   12662: 'Pump6: Pressure recording: warning, value undershot', class Pump Warning Alarm, trigger "Pump6_Pressure_Record_DBW_142" bit 10
   12663: 'Pump6: Pressure recording: fault, value exceeded', class Pump Error Alarm, trigger "Pump6_Pressure_Record_DBW_142" bit 11
   12664: 'Pump6: Pressure recording: fault, value undershot', class Pump Error Alarm, trigger "Pump6_Pressure_Record_DBW_142" bit 12
   12665: 'Pump6: Temp. recording HP heat exch.: measured value outside measuring range', class Pump Warning Alarm, trigger "Pump6_Heatexchanger_DBW_220" bit 8
   12666: 'Pump6: Temp. recording HP heat exch.: warning, value exceeded', class Pump Warning Alarm, trigger "Pump6_Heatexchanger_DBW_220" bit 9
   12667: 'Pump6: Temp. recording HP heat exch.: warning, value undershot', class Pump Warning Alarm, trigger "Pump6_Heatexchanger_DBW_220" bit 10
   12668: 'Pump6: Temp. recording HP heat exch.: fault, value exceeded', class Pump Error Alarm, trigger "Pump6_Heatexchanger_DBW_220" bit 11
   12669: 'Pump6: Temp. recording HP heat exch.: fault, value undershot', class Pump Error Alarm, trigger "Pump6_Heatexchanger_DBW_220" bit 12
   10101: 'Mixinghead hydraulic: Motor protection switch has tripped', class Mixing Hydraulic Errors, trigger "Mixinghead_Hydraulic_DBW2" bit 8
   10102: 'Mixinghead hydraulic: Min. fill level hydraulic oil undershot', class Mixing Hydraulic Errors, trigger "Mixinghead_Hydraulic_DBW2" bit 9
   10103: 'Mixinghead hydraulic: Warning max. temperature exceeded', class Mixing Hydraulic Warning, trigger "Mixinghead_Hydraulic_DBW2" bit 10
   10104: 'Mixinghead hydraulic: HP filter contaminated', class Mixing Hydraulic Warning, trigger "Mixinghead_Hydraulic_DBW2" bit 11
   10105: 'Mixinghead hydraulic: Activation max. temperature exceeded', class Mixing Hydraulic Errors, trigger "Mixinghead_Hydraulic_DBW2" bit 12
   10106: 'Mixinghead hydraulic: Return filter contaminated', class Mixing Hydraulic Warning, trigger "Mixinghead_Hydraulic_DBW2" bit 13
   10107: 'Mixinghead hydraulic: Cable break at pressure switch', class Mixing Hydraulic Errors, trigger "Mixinghead_Hydraulic_DBW2" bit 14
   10108: 'Mixinghead hydraulic: Max. pressure not reached', class Mixing Hydraulic Errors, trigger "Mixinghead_Hydraulic_DBW2" bit 15
   10109: 'Mixinghead hydraulic: Moog filter contaminated', class Mixing Hydraulic Warning, trigger "Mixinghead_Hydraulic_DBW2" bit 0
   10110: 'Mixinghead hydraulic: Min. fill level filter pump', class Mixing Hydraulic Warning, trigger "Mixinghead_Hydraulic_DBW2" bit 1
   10111: 'Mixinghead hydraulic: Motor protecting switch of filter pump tripped', class Mixing Hydraulic Errors, trigger "Mixinghead_Hydraulic_DBW2" bit 2
   10112: 'Mixinghead hydraulic: Max. fill level filter pump', class Mixing Hydraulic Errors, trigger "Mixinghead_Hydraulic_DBW2" bit 3
   10113: 'Mixinghead hydraulic: Filter bypass fault', class Mixing Hydraulic Warning, trigger "Mixinghead_Hydraulic_DBW2" bit 4
   10114: 'Mixinghead hydraulic:', class Mixing Hydraulic Warning, trigger "Mixinghead_Hydraulic_DBW2" bit 5
   10115: 'Mixinghead hydraulic:', class Mixing Hydraulic Errors, trigger "Mixinghead_Hydraulic_DBW2" bit 6
   10116: 'Mixinghead hydraulic:', class Mixing Hydraulic Errors, trigger "Mixinghead_Hydraulic_DBW2" bit 7
   15001: 'Mixinghead 01: Mixinghead does not open', class Mixing Head Errors, trigger "Mixinghead_MHControl1_DBW_2" bit 8
   15002: 'Mixinghead 01: Mixinghead does not close', class Mixing Head Errors, trigger "Mixinghead_MHControl1_DBW_2" bit 9
   15003: 'Mixinghead 01: Entry cancelled', class Mixing Head Warning, trigger "Mixinghead_MHControl1_DBW_2" bit 10
   15004: 'Mixinghead 01: Mixinghead open without activation', class Mixing Head Errors, trigger "Mixinghead_MHControl1_DBW_2" bit 11
   15005: 'Mixinghead 01: Mixinghead close during entry', class Mixing Head Warning, trigger "Mixinghead_MHControl1_DBW_2" bit 12
   15006: 'Mixinghead 01: Warning, shot time too short', class Mixing Head Warning, trigger "Mixinghead_MHControl1_DBW_2" bit 13
   15007: 'Mixinghead 01: Warning , shot time too long', class Mixing Head Warning, trigger "Mixinghead_MHControl1_DBW_2" bit 14
   15008: 'Mixinghead 01: Fault, shot time too short', class Mixing Head Warning, trigger "Mixinghead_MHControl1_DBW_2" bit 15
   15009: 'Mixinghead 01: Mixinghead collides when opening or closing', class Mixing Head Warning, trigger "Mixinghead_MHControl1_DBW_2" bit 0
   15010: 'Mixinghead 01: Runtime monitoring when locking mixing head', class Mixing Head Warning, trigger "Mixinghead_MHControl1_DBW_2" bit 1
   15011: 'Mixinghead 01: Runtime monitoring when unlocking mixing head', class Mixing Head Warning, trigger "Mixinghead_MHControl1_DBW_2" bit 2
   15012: 'Mixinghead 01:', class Mixing Head Warning, trigger "Mixinghead_MHControl1_DBW_2" bit 3
   15013: 'Mixinghead 01: Min. Pressure for the cleaning air', class Mixing Head Warning, trigger "Mixinghead_MHControl1_DBW_2" bit 4
   15014: 'Mixinghead 01: Max. Pressure for the cleaning air', class Mixing Head Warning, trigger "Mixinghead_MHControl1_DBW_2" bit 5
   15015: 'Mixinghead 01:', class Mixing Head Warning, trigger "Mixinghead_MHControl1_DBW_2" bit 6
   15016: 'Mixinghead 01: Component required in entry is not enabled at this mixing head', class Mixing Head Errors, trigger "Mixinghead_MHControl1_DBW_2" bit 7
   15017: 'Mixinghead 01: Cleaning piston: Moving out too slow', class Mixing Head Errors, trigger "Mixinghead_Cpiston1_DBW_34" bit 8
   15018: 'Mixinghead 01: Cleaning piston: Moving in too slow', class Mixing Head Errors, trigger "Mixinghead_Cpiston1_DBW_34" bit 9
   15019: 'Mixinghead 01: Cleaning piston: Proximity switch defect', class Mixinghead Error Archive Foaming, trigger "Mixinghead_Cpiston1_DBW_34" bit 10
   15020: 'Mixinghead 01: Cleaning piston: Leaves its home position in entry', class Mixing Head Errors, trigger "Mixinghead_Cpiston1_DBW_34" bit 11
   15021: 'Mixinghead 01: Cleaning piston: Not defined', class Mixing Head Warning, trigger "Mixinghead_Cpiston1_DBW_34" bit 12
   15022: 'Mixinghead 01: Cleaning piston:', class Mixing Head Warning, trigger "Mixinghead_Cpiston1_DBW_34" bit 13
   15023: 'Mixinghead 01: Cleaning piston:', class Mixing Head Warning, trigger "Mixinghead_Cpiston1_DBW_34" bit 14
   15024: 'Mixinghead 01: Cleaning piston:', class Mixing Head Warning, trigger "Mixinghead_Cpiston1_DBW_34" bit 15
   15025: 'Mixinghead 01: Cleaning piston: Controller at upper limit', class Mixing Head Warning, trigger "Mixinghead_Cpiston1_DBW_34" bit 0
   15026: 'Mixinghead 01: Cleaning piston: Controller at lower limit', class Mixing Head Warning, trigger "Mixinghead_Cpiston1_DBW_34" bit 1
   15027: 'Mixinghead 01: Cleaning piston:', class Mixing Head Warning, trigger "Mixinghead_Cpiston1_DBW_34" bit 2
   15028: 'Mixinghead 01: Cleaning piston: Front position not reached', class Mixing Head Warning, trigger "Mixinghead_Cpiston1_DBW_34" bit 3
   15029: 'Mixinghead 01: Cleaning piston: Rear position not reached', class Mixing Head Warning, trigger "Mixinghead_Cpiston1_DBW_34" bit 4
   15030: 'Mixinghead 01: Cleaning piston: Home position not reached', class Mixing Head Warning, trigger "Mixinghead_Cpiston1_DBW_34" bit 5
   15031: 'Mixinghead 01: Cleaning piston:', class Mixing Head Warning, trigger "Mixinghead_Cpiston1_DBW_34" bit 6
   15032: 'Mixinghead 01: Cleaning piston:', class Mixing Head Warning, trigger "Mixinghead_Cpiston1_DBW_34" bit 7
   15040: 'Mixinghead 01: Connection 01: Temperature recording: Measuring value outside measuring range', class Mixinghead Warn Archv Foam, trigger "Mixinghead_Temperature_MH1_Con1_DBW70" bit 8
   15041: 'Mixinghead 01: Connection 01: Temperature recording: Warning, value exceeded', class Mixing Head Warning, trigger "Mixinghead_Temperature_MH1_Con1_DBW70" bit 9
   15042: 'Mixinghead 01: Connection 01: Temperature recording: Warning, value undershot', class Mixing Head Warning, trigger "Mixinghead_Temperature_MH1_Con1_DBW70" bit 10
   15043: 'Mixinghead 01: Connection 01: Temperature recording: Fault, value exceeded', class Mixing Head Errors, trigger "Mixinghead_Temperature_MH1_Con1_DBW70" bit 11
   15044: 'Mixinghead 01: Connection 01: Temperature recording: Fault, value undershot', class Mixing Head Errors, trigger "Mixinghead_Temperature_MH1_Con1_DBW70" bit 12
   15045: 'Mixinghead 01: Connection 02: Temperature recording: Measuring value outside measuring range', class Mixinghead Warn Archv Foam, trigger "Mixinghead_Temperature_MH1_Con2_DBW104" bit 8
   15046: 'Mixinghead 01: Connection 02: Temperature recording: Warning, value exceeded', class Mixing Head Warning, trigger "Mixinghead_Temperature_MH1_Con2_DBW104" bit 9
   15047: 'Mixinghead 01: Connection 02: Temperature recording: Warning, value undershot', class Mixing Head Warning, trigger "Mixinghead_Temperature_MH1_Con2_DBW104" bit 10
   15048: 'Mixinghead 01: Connection 02: Temperature recording: Fault, value exceeded', class Mixing Head Errors, trigger "Mixinghead_Temperature_MH1_Con2_DBW104" bit 11
   15049: 'Mixinghead 01: Connection 02: Temperature recording: Fault, value undershot', class Mixing Head Errors, trigger "Mixinghead_Temperature_MH1_Con2_DBW104" bit 12
   15050: 'Mixinghead 01: Connection 03: Temperature recording: Measuring value outside measuring range', class Mixing Head Warning, trigger "Mixinghead_Temperature_MH1_Con3_DBW138" bit 8
   15051: 'Mixinghead 01: Connection 03: Temperature recording: Warning, value exceeded', class Mixing Head Warning, trigger "Mixinghead_Temperature_MH1_Con3_DBW138" bit 9
   15052: 'Mixinghead 01: Connection 03: Temperature recording: Warning, value undershot', class Mixing Head Warning, trigger "Mixinghead_Temperature_MH1_Con3_DBW138" bit 10
   15053: 'Mixinghead 01: Connection 03: Temperature recording: Fault, value exceeded', class Mixing Head Errors, trigger "Mixinghead_Temperature_MH1_Con3_DBW138" bit 11
   15054: 'Mixinghead 01: Connection 03: Temperature recording: Fault, value undershot', class Mixing Head Errors, trigger "Mixinghead_Temperature_MH1_Con3_DBW138" bit 12
   15055: 'Mixinghead 01: Connection 04: Temperature recording: Measuring value outside measuring range', class Mixing Head Warning, trigger "Mixinghead_Temperature_MH1_Con4_DBW172" bit 8
   15056: 'Mixinghead 01: Connection 04: Temperature recording: Warning, value exceeded', class Mixing Head Warning, trigger "Mixinghead_Temperature_MH1_Con4_DBW172" bit 9
   15057: 'Mixinghead 01: Connection 04: Temperature recording: Warning, value undershot', class Mixing Head Warning, trigger "Mixinghead_Temperature_MH1_Con4_DBW172" bit 10
   15058: 'Mixinghead 01: Connection 04: Temperature recording: Fault, value exceeded', class Mixing Head Errors, trigger "Mixinghead_Temperature_MH1_Con4_DBW172" bit 11
   15059: 'Mixinghead 01: Connection 04: Temperature recording: Fault, value undershot', class Mixing Head Errors, trigger "Mixinghead_Temperature_MH1_Con4_DBW172" bit 12
   15060: 'Mixinghead 01: Connection 05: Temperature recording: Measuring value outside measuring range', class Mixing Head Warning, trigger "Mixinghead_Temperature_MH1_Con5_DBW206" bit 8
   15061: 'Mixinghead 01: Connection 05: Temperature recording: Warning, value exceeded', class Mixing Head Warning, trigger "Mixinghead_Temperature_MH1_Con5_DBW206" bit 9
   15062: 'Mixinghead 01: Connection 05: Temperature recording: Warning, value undershot', class Mixing Head Warning, trigger "Mixinghead_Temperature_MH1_Con5_DBW206" bit 10
   15063: 'Mixinghead 01: Connection 05: Temperature recording: Fault, value exceeded', class Mixing Head Errors, trigger "Mixinghead_Temperature_MH1_Con5_DBW206" bit 11
   15064: 'Mixinghead 01: Connection 05: Temperature recording: Fault, value undershot', class Mixing Head Errors, trigger "Mixinghead_Temperature_MH1_Con5_DBW206" bit 12
   15065: 'Mixinghead 01: Connection 06: Temperature recording: Measuring value outside measuring range', class Mixing Head Warning, trigger "Mixinghead_Temperature_MH1_Con6_DBW240" bit 8
   15066: 'Mixinghead 01: Connection 06: Temperature recording: Warning, value exceeded', class Mixing Head Warning, trigger "Mixinghead_Temperature_MH1_Con6_DBW240" bit 9
   15067: 'Mixinghead 01: Connection 06: Temperature recording: Warning, value undershot', class Mixing Head Warning, trigger "Mixinghead_Temperature_MH1_Con6_DBW240" bit 10
   15068: 'Mixinghead 01: Connection 06: Temperature recording: Fault, value exceeded', class Mixing Head Errors, trigger "Mixinghead_Temperature_MH1_Con6_DBW240" bit 11
   15069: 'Mixinghead 01: Connection 06: Temperature recording: Fault, value undershot', class Mixing Head Errors, trigger "Mixinghead_Temperature_MH1_Con6_DBW240" bit 12
   15070: 'Mixinghead 01: Connection 01: Pressure recording: Measuring value outside measuring range', class Mixing Head Warning, trigger "Mixinghead_Pressure_MH1_Con1_DBW274" bit 8
   15071: 'Mixinghead 01: Connection 01: Pressure recording: Warning, value exceeded', class Mixing Head Warning, trigger "Mixinghead_Pressure_MH1_Con1_DBW274" bit 9
   15072: 'Mixinghead 01: Connection 01: Pressure recording: Warning, value undershot', class Mixing Head Warning, trigger "Mixinghead_Pressure_MH1_Con1_DBW274" bit 10
   15073: 'Mixinghead 01: Connection 01: Pressure recording: Fault, value exceeded', class Mixing Head Errors, trigger "Mixinghead_Pressure_MH1_Con1_DBW274" bit 11
   15075: 'Mixinghead 01: Connection 02: Pressure recording: Measuring value outside measuring range', class Mixing Head Warning, trigger "Mixinghead_Pressure_MH1_Con2_DBW308" bit 8
   15076: 'Mixinghead 01: Connection 02: Pressure recording: Warning, value exceeded', class Mixing Head Warning, trigger "Mixinghead_Pressure_MH1_Con2_DBW308" bit 9
   15077: 'Mixinghead 01: Connection 02: Pressure recording: Warning, value undershot', class Mixing Head Warning, trigger "Mixinghead_Pressure_MH1_Con2_DBW308" bit 10
   15078: 'Mixinghead 01: Connection 02: Pressure recording: Fault, value exceeded', class Mixing Head Errors, trigger "Mixinghead_Pressure_MH1_Con2_DBW308" bit 11
   15079: 'Mixinghead 01: Connection 02: Pressure recording: Fault, value undershot', class Mixing Head Errors, trigger "Mixinghead_Pressure_MH1_Con2_DBW308" bit 12
   15080: 'Mixinghead 01: Connection 03: Pressure recording: Measuring value outside measuring range', class Mixing Head Warning, trigger "Mixinghead_Pressure_MH1_Con3_DBW342" bit 8
   15081: 'Mixinghead 01: Connection 03: Pressure recording: Warning, value exceeded', class Mixing Head Warning, trigger "Mixinghead_Pressure_MH1_Con3_DBW342" bit 9
   15082: 'Mixinghead 01: Connection 03: Pressure recording: Warning, value undershot', class Mixing Head Warning, trigger "Mixinghead_Pressure_MH1_Con3_DBW342" bit 10
   15083: 'Mixinghead 01: Connection 03: Pressure recording: Fault, value exceeded', class Mixing Head Errors, trigger "Mixinghead_Pressure_MH1_Con3_DBW342" bit 11
   15084: 'Mixinghead 01: Connection 03: Pressure recording: Fault, value undershot', class Mixing Head Errors, trigger "Mixinghead_Pressure_MH1_Con3_DBW342" bit 12
   15085: 'Mixinghead 01: Connection 04: Pressure recording: Measuring value outside measuring range', class Mixing Head Warning, trigger "Mixinghead_Pressure_MH1_Con4_DBW376" bit 8
   15086: 'Mixinghead 01: Connection 04: Pressure recording: Warning, value exceeded', class Mixing Head Warning, trigger "Mixinghead_Pressure_MH1_Con4_DBW376" bit 9
   15087: 'Mixinghead 01: Connection 04: Pressure recording: Warning, value undershot', class Mixing Head Warning, trigger "Mixinghead_Pressure_MH1_Con4_DBW376" bit 10
   15088: 'Mixinghead 01: Connection 04: Pressure recording: Fault, value exceeded', class Mixing Head Errors, trigger "Mixinghead_Pressure_MH1_Con4_DBW376" bit 11
   15089: 'Mixinghead 01: Connection 04: Pressure recording: Fault, value undershot', class Mixing Head Errors, trigger "Mixinghead_Pressure_MH1_Con4_DBW376" bit 12
   15090: 'Mixinghead 01: Connection 05: Pressure recording: Measuring value outside measuring range', class Mixing Head Warning, trigger "Mixinghead_Pressure_MH1_Con5_DBW410" bit 8
   15091: 'Mixinghead 01: Connection 05: Pressure recording: Warning, value exceeded', class Mixing Head Warning, trigger "Mixinghead_Pressure_MH1_Con5_DBW410" bit 9
   15092: 'Mixinghead 01: Connection 05: Pressure recording: Warning, value undershot', class Mixing Head Warning, trigger "Mixinghead_Pressure_MH1_Con5_DBW410" bit 10
   15093: 'Mixinghead 01: Connection 05: Pressure recording: Fault, value exceeded', class Mixing Head Errors, trigger "Mixinghead_Pressure_MH1_Con5_DBW410" bit 11
   15094: 'Mixinghead 01: Connection 05: Pressure recording: Fault, value undershot', class Mixing Head Errors, trigger "Mixinghead_Pressure_MH1_Con5_DBW410" bit 12
   15095: 'Mixinghead 01: Connection 06: Pressure recording: Measuring value outside measuring range', class Mixing Head Warning, trigger "Mixinghead_Pressure_MH1_Con6_DBW444" bit 8
   15096: 'Mixinghead 01: Connection 06: Pressure recording: Warning, value exceeded', class Mixing Head Warning, trigger "Mixinghead_Pressure_MH1_Con6_DBW444" bit 9
   15097: 'Mixinghead 01: Connection 06: Pressure recording: Warning, value undershot', class Mixing Head Warning, trigger "Mixinghead_Pressure_MH1_Con6_DBW444" bit 10
   15098: 'Mixinghead 01: Connection 06: Pressure recording: Fault, value exceeded', class Mixing Head Errors, trigger "Mixinghead_Pressure_MH1_Con6_DBW444" bit 11
   15099: 'Mixinghead 01: Connection 06: Pressure recording: Fault, value undershot', class Mixing Head Errors, trigger "Mixinghead_Pressure_MH1_Con6_DBW444" bit 12
   15074: 'Mixinghead 01: Connection 01: Pressure recording: Fault, value undershot', class Mixing Head Errors, trigger "Mixinghead_Pressure_MH1_Con1_DBW274" bit 12
   15101: 'Mixinghead 02: Mixinghead does not open', class Mixing Head Errors, trigger "Mixinghead_MHControl2_DBW_4" bit 8
   15102: 'Mixinghead 02: Mixinghead does not close', class Mixing Head Errors, trigger "Mixinghead_MHControl2_DBW_4" bit 9
   15103: 'Mixinghead 02: Entry cancelled', class Mixing Head Warning, trigger "Mixinghead_MHControl2_DBW_4" bit 10
   15104: 'Mixinghead 02: Mixinghead open without activation', class Mixing Head Errors, trigger "Mixinghead_MHControl2_DBW_4" bit 11
   15105: 'Mixinghead 02: Mixinghead close during entry', class Mixing Head Warning, trigger "Mixinghead_MHControl2_DBW_4" bit 12
   15106: 'Mixinghead 02: Warning, shot time too short', class Mixing Head Warning, trigger "Mixinghead_MHControl2_DBW_4" bit 13
   15107: 'Mixinghead 02: Warning , shot time too long', class Mixing Head Warning, trigger "Mixinghead_MHControl2_DBW_4" bit 14
   15108: 'Mixinghead 02: Fault, shot time too short', class Mixing Head Warning, trigger "Mixinghead_MHControl2_DBW_4" bit 15
   15109: 'Mixinghead 02: Mixinghead collides when opening or closing', class Mixing Head Warning, trigger "Mixinghead_MHControl2_DBW_4" bit 0
   15110: 'Mixinghead 02: Runtime monitoring when locking mixing head', class Mixing Head Warning, trigger "Mixinghead_MHControl2_DBW_4" bit 1
   15111: 'Mixinghead 02: Runtime monitoring when unlocking mixing head', class Mixing Head Warning, trigger "Mixinghead_MHControl2_DBW_4" bit 2
   15112: 'Mixinghead 02:', class Mixing Head Warning, trigger "Mixinghead_MHControl2_DBW_4" bit 3
   15113: 'Mixinghead 02:', class Mixing Head Warning, trigger "Mixinghead_MHControl2_DBW_4" bit 4
   15114: 'Mixinghead 02:', class Mixing Head Warning, trigger "Mixinghead_MHControl2_DBW_4" bit 5
   15115: 'Mixinghead 02:', class Mixing Head Warning, trigger "Mixinghead_MHControl2_DBW_4" bit 6
   15116: 'Mixinghead 02: Component required in entry is not enabled at this mixing head', class Mixing Head Errors, trigger "Mixinghead_MHControl2_DBW_4" bit 7
   15117: 'Mixinghead 02: Cleaning piston: Moving out too slow', class Mixing Head Errors, trigger "Mixinghead_Cpiston2_DBW_36" bit 8
   15118: 'Mixinghead 02: Cleaning piston: Moving in too slow', class Mixing Head Errors, trigger "Mixinghead_Cpiston2_DBW_36" bit 9
   15119: 'Mixinghead 02: Cleaning piston: Proximity switch defect', class Mixing Head Errors, trigger "Mixinghead_Cpiston2_DBW_36" bit 10
   15120: 'Mixinghead 02: Cleaning piston: Leaves its home position in entry', class Mixing Head Errors, trigger "Mixinghead_Cpiston2_DBW_36" bit 11
   15121: 'Mixinghead 02: Cleaning piston: Not defined', class Mixing Head Warning, trigger "Mixinghead_Cpiston2_DBW_36" bit 12
   15122: 'Mixinghead 02: Cleaning piston:', class Mixing Head Warning, trigger "Mixinghead_Cpiston2_DBW_36" bit 13
   15123: 'Mixinghead 02: Cleaning piston:', class Mixing Head Warning, trigger "Mixinghead_Cpiston2_DBW_36" bit 14
   15124: 'Mixinghead 02: Cleaning piston:', class Mixing Head Warning, trigger "Mixinghead_Cpiston2_DBW_36" bit 15
   15125: 'Mixinghead 02: Cleaning piston: Controller at upper limit', class Mixing Head Warning, trigger "Mixinghead_Cpiston2_DBW_36" bit 0
   15126: 'Mixinghead 02: Cleaning piston: Controller at lower limit', class Mixing Head Warning, trigger "Mixinghead_Cpiston2_DBW_36" bit 1
   15127: 'Mixinghead 02: Cleaning piston:', class Mixing Head Warning, trigger "Mixinghead_Cpiston2_DBW_36" bit 2
   15128: 'Mixinghead 02: Cleaning piston: Front position not reached', class Mixing Head Warning, trigger "Mixinghead_Cpiston2_DBW_36" bit 3
   15129: 'Mixinghead 02: Cleaning piston: Rear position not reached', class Mixing Head Warning, trigger "Mixinghead_Cpiston2_DBW_36" bit 4
   15130: 'Mixinghead 02: Cleaning piston: Home position not reached', class Mixing Head Warning, trigger "Mixinghead_Cpiston2_DBW_36" bit 5
   15131: 'Mixinghead 02: Cleaning piston:', class Mixing Head Warning, trigger "Mixinghead_Cpiston2_DBW_36" bit 6
   15132: 'Mixinghead 02: Cleaning piston:', class Mixing Head Warning, trigger "Mixinghead_Cpiston2_DBW_36" bit 7
   15140: 'Mixinghead 02: Connection 01: Temperature recording: Measuring value outside measuring range', class Mixing Head Warning, trigger "Mixinghead_Temperature_MH2_Con1_DBW72" bit 8
   15141: 'Mixinghead 02: Connection 01: Temperature recording: Warning, value exceeded', class Mixing Head Warning, trigger "Mixinghead_Temperature_MH2_Con1_DBW72" bit 9
   15142: 'Mixinghead 02: Connection 01: Temperature recording: Warning, value undershot', class Mixing Head Warning, trigger "Mixinghead_Temperature_MH2_Con1_DBW72" bit 10
   15143: 'Mixinghead 02: Connection 01: Temperature recording: Fault, value exceeded', class Mixing Head Errors, trigger "Mixinghead_Temperature_MH2_Con1_DBW72" bit 11
   15144: 'Mixinghead 02: Connection 01: Temperature recording: Fault, value undershot', class Mixing Head Errors, trigger "Mixinghead_Temperature_MH2_Con1_DBW72" bit 12
   15145: 'Mixinghead 02: Connection 02: Temperature recording: Measuring value outside measuring range', class Mixing Head Warning, trigger "Mixinghead_Temperature_MH2_Con2_DBW106" bit 8
   15146: 'Mixinghead 02: Connection 02: Temperature recording: Warning, value exceeded', class Mixing Head Warning, trigger "Mixinghead_Temperature_MH2_Con2_DBW106" bit 9
   15147: 'Mixinghead 02: Connection 02: Temperature recording: Warning, value undershot', class Mixing Head Warning, trigger "Mixinghead_Temperature_MH2_Con2_DBW106" bit 10
   15148: 'Mixinghead 02: Connection 02: Temperature recording: Fault, value exceeded', class Mixing Head Errors, trigger "Mixinghead_Temperature_MH2_Con2_DBW106" bit 11
   15149: 'Mixinghead 02: Connection 02: Temperature recording: Fault, value undershot', class Mixing Head Errors, trigger "Mixinghead_Temperature_MH2_Con2_DBW106" bit 12
   15150: 'Mixinghead 02: Connection 03: Temperature recording: Measuring value outside measuring range', class Mixing Head Warning, trigger "Mixinghead_Temperature_MH2_Con3_DBW140" bit 8
   15151: 'Mixinghead 02: Connection 03: Temperature recording: Warning, value exceeded', class Mixing Head Warning, trigger "Mixinghead_Temperature_MH2_Con3_DBW140" bit 9
   15152: 'Mixinghead 02: Connection 03: Temperature recording: Warning, value undershot', class Mixing Head Warning, trigger "Mixinghead_Temperature_MH2_Con3_DBW140" bit 10
   15153: 'Mixinghead 02: Connection 03: Temperature recording: Fault, value exceeded', class Mixing Head Errors, trigger "Mixinghead_Temperature_MH2_Con3_DBW140" bit 11
   15154: 'Mixinghead 02: Connection 03: Temperature recording: Fault, value undershot', class Mixing Head Errors, trigger "Mixinghead_Temperature_MH2_Con3_DBW140" bit 12
   15155: 'Mixinghead 02: Connection 04: Temperature recording: Measuring value outside measuring range', class Mixing Head Warning, trigger "Mixinghead_Temperature_MH2_Con4_DBW174" bit 8
   15156: 'Mixinghead 02: Connection 04: Temperature recording: Warning, value exceeded', class Mixing Head Warning, trigger "Mixinghead_Temperature_MH2_Con4_DBW174" bit 9
   15157: 'Mixinghead 02: Connection 04: Temperature recording: Warning, value undershot', class Mixing Head Warning, trigger "Mixinghead_Temperature_MH2_Con4_DBW174" bit 10
   15158: 'Mixinghead 02: Connection 04: Temperature recording: Fault, value exceeded', class Mixing Head Errors, trigger "Mixinghead_Temperature_MH2_Con4_DBW174" bit 11
   15159: 'Mixinghead 02: Connection 04: Temperature recording: Fault, value undershot', class Mixing Head Errors, trigger "Mixinghead_Temperature_MH2_Con4_DBW174" bit 12
   15160: 'Mixinghead 02: Connection 05: Temperature recording: Measuring value outside measuring range', class Mixing Head Warning, trigger "Mixinghead_Temperature_MH2_Con5_DBW208" bit 8
   15161: 'Mixinghead 02: Connection 05: Temperature recording: Warning, value exceeded', class Mixing Head Warning, trigger "Mixinghead_Temperature_MH2_Con5_DBW208" bit 9
   15162: 'Mixinghead 02: Connection 05: Temperature recording: Warning, value undershot', class Mixing Head Warning, trigger "Mixinghead_Temperature_MH2_Con5_DBW208" bit 10
   15163: 'Mixinghead 02: Connection 05: Temperature recording: Fault, value exceeded', class Mixing Head Errors, trigger "Mixinghead_Temperature_MH2_Con5_DBW208" bit 11
   15164: 'Mixinghead 02: Connection 05: Temperature recording: Fault, value undershot', class Mixing Head Errors, trigger "Mixinghead_Temperature_MH2_Con5_DBW208" bit 12
   15165: 'Mixinghead 02: Connection 06: Temperature recording: Measuring value outside measuring range', class Mixing Head Warning, trigger "Mixinghead_Temperature_MH2_Con6_DBW242" bit 8
   15166: 'Mixinghead 02: Connection 06: Temperature recording: Warning, value exceeded', class Mixing Head Warning, trigger "Mixinghead_Temperature_MH2_Con6_DBW242" bit 9
   15167: 'Mixinghead 02: Connection 06: Temperature recording: Warning, value undershot', class Mixing Head Warning, trigger "Mixinghead_Temperature_MH2_Con6_DBW242" bit 10
   15168: 'Mixinghead 02: Connection 06: Temperature recording: Fault, value exceeded', class Mixing Head Errors, trigger "Mixinghead_Temperature_MH2_Con6_DBW242" bit 11
   15169: 'Mixinghead 02: Connection 06: Temperature recording: Fault, value undershot', class Mixing Head Errors, trigger "Mixinghead_Temperature_MH2_Con6_DBW242" bit 12
   15170: 'Mixinghead 02: Connection 01: Pressure recording: Measuring value outside measuring range', class Mixing Head Warning, trigger "Mixinghead_Pressure_MH2_Con1_DBW276" bit 8
   15171: 'Mixinghead 02: Connection 01: Pressure recording: Warning, value exceeded', class Mixing Head Warning, trigger "Mixinghead_Pressure_MH2_Con1_DBW276" bit 9
   15172: 'Mixinghead 02: Connection 01: Pressure recording: Warning, value undershot', class Mixing Head Warning, trigger "Mixinghead_Pressure_MH2_Con1_DBW276" bit 10
   15173: 'Mixinghead 02: Connection 01: Pressure recording: Fault, value exceeded', class Mixing Head Errors, trigger "Mixinghead_Pressure_MH2_Con1_DBW276" bit 11
   15174: 'Mixinghead 02: Connection 01: Pressure recording: Fault, value undershot', class Mixing Head Errors, trigger "Mixinghead_Pressure_MH2_Con1_DBW276" bit 12
   15175: 'Mixinghead 02: Connection 02: Pressure recording: Measuring value outside measuring range', class Mixing Head Warning, trigger "Mixinghead_Pressure_MH2_Con2_DBW310" bit 8
   15176: 'Mixinghead 02: Connection 02: Pressure recording: Warning, value exceeded', class Mixing Head Warning, trigger "Mixinghead_Pressure_MH2_Con2_DBW310" bit 9
   15177: 'Mixinghead 02: Connection 02: Pressure recording: Warning, value undershot', class Mixing Head Warning, trigger "Mixinghead_Pressure_MH2_Con2_DBW310" bit 10
   15178: 'Mixinghead 02: Connection 02: Pressure recording: Fault, value exceeded', class Mixing Head Errors, trigger "Mixinghead_Pressure_MH2_Con2_DBW310" bit 11
   15179: 'Mixinghead 02: Connection 02: Pressure recording: Fault, value undershot', class Mixing Head Errors, trigger "Mixinghead_Pressure_MH2_Con2_DBW310" bit 12
   15180: 'Mixinghead 02: Connection 03: Pressure recording: Measuring value outside measuring range', class Mixing Head Warning, trigger "Mixinghead_Pressure_MH2_Con3_DBW344" bit 8
   15181: 'Mixinghead 02: Connection 03: Pressure recording: Warning, value exceeded', class Mixing Head Warning, trigger "Mixinghead_Pressure_MH2_Con3_DBW344" bit 9
   15182: 'Mixinghead 02: Connection 03: Pressure recording: Warning, value undershot', class Mixing Head Warning, trigger "Mixinghead_Pressure_MH2_Con3_DBW344" bit 10
   15183: 'Mixinghead 02: Connection 03: Pressure recording: Fault, value exceeded', class Mixing Head Errors, trigger "Mixinghead_Pressure_MH2_Con3_DBW344" bit 11
   15184: 'Mixinghead 02: Connection 03: Pressure recording: Fault, value undershot', class Mixing Head Errors, trigger "Mixinghead_Pressure_MH2_Con3_DBW344" bit 12
   15185: 'Mixinghead 02: Connection 04: Pressure recording: Measuring value outside measuring range', class Mixing Head Warning, trigger "Mixinghead_Pressure_MH2_Con4_DBW378" bit 8
   15186: 'Mixinghead 02: Connection 04: Pressure recording: Warning, value exceeded', class Mixing Head Warning, trigger "Mixinghead_Pressure_MH2_Con4_DBW378" bit 9
   15187: 'Mixinghead 02: Connection 04: Pressure recording: Warning, value undershot', class Mixing Head Warning, trigger "Mixinghead_Pressure_MH2_Con4_DBW378" bit 10
   15188: 'Mixinghead 02: Connection 04: Pressure recording: Fault, value exceeded', class Mixing Head Errors, trigger "Mixinghead_Pressure_MH2_Con4_DBW378" bit 11
   15189: 'Mixinghead 02: Connection 04: Pressure recording: Fault, value undershot', class Mixing Head Errors, trigger "Mixinghead_Pressure_MH2_Con4_DBW378" bit 12
   15190: 'Mixinghead 02: Connection 05: Pressure recording: Measuring value outside measuring range', class Mixing Head Warning, trigger "Mixinghead_Pressure_MH2_Con5_DBW412" bit 8
   15191: 'Mixinghead 02: Connection 05: Pressure recording: Warning, value exceeded', class Mixing Head Warning, trigger "Mixinghead_Pressure_MH2_Con5_DBW412" bit 9
   15192: 'Mixinghead 02: Connection 05: Pressure recording: Warning, value undershot', class Mixing Head Warning, trigger "Mixinghead_Pressure_MH2_Con5_DBW412" bit 10
   15193: 'Mixinghead 02: Connection 05: Pressure recording: Fault, value exceeded', class Mixing Head Errors, trigger "Mixinghead_Pressure_MH2_Con5_DBW412" bit 11
   15194: 'Mixinghead 02: Connection 05: Pressure recording: Fault, value undershot', class Mixing Head Errors, trigger "Mixinghead_Pressure_MH2_Con5_DBW412" bit 12
   15195: 'Mixinghead 02: Connection 06: Pressure recording: Measuring value outside measuring range', class Mixing Head Warning, trigger "Mixinghead_Pressure_MH2_Con6_DBW446" bit 8
   15196: 'Mixinghead 02: Connection 06: Pressure recording: Warning, value exceeded', class Mixing Head Warning, trigger "Mixinghead_Pressure_MH2_Con6_DBW446" bit 9
   15197: 'Mixinghead 02: Connection 06: Pressure recording: Warning, value undershot', class Mixing Head Warning, trigger "Mixinghead_Pressure_MH2_Con6_DBW446" bit 10
   15198: 'Mixinghead 02: Connection 06: Pressure recording: Fault, value exceeded', class Mixing Head Errors, trigger "Mixinghead_Pressure_MH2_Con6_DBW446" bit 11
   15199: 'Mixinghead 02: Connection 06: Pressure recording: Fault, value undershot', class Mixing Head Errors, trigger "Mixinghead_Pressure_MH2_Con6_DBW446" bit 12
   15201: 'Mixinghead 03: Mixinghead does not open', class Mixing Head Errors, trigger "Mixinghead_MHControl3_DBW_6" bit 8
   15202: 'Mixinghead 03: Mixinghead does not close', class Mixing Head Errors, trigger "Mixinghead_MHControl3_DBW_6" bit 9
   15203: 'Mixinghead 03: Entry cancelled', class Mixing Head Warning, trigger "Mixinghead_MHControl3_DBW_6" bit 10
   15204: 'Mixinghead 03: Mixinghead open without activation', class Mixing Head Errors, trigger "Mixinghead_MHControl3_DBW_6" bit 11
   15205: 'Mixinghead 03: Mixinghead close during entry', class Mixing Head Warning, trigger "Mixinghead_MHControl3_DBW_6" bit 12
   15206: 'Mixinghead 03: Warning, shot time too short', class Mixing Head Warning, trigger "Mixinghead_MHControl3_DBW_6" bit 13
   15207: 'Mixinghead 03: Warning , shot time too long', class Mixing Head Warning, trigger "Mixinghead_MHControl3_DBW_6" bit 14
   15208: 'Mixinghead 03: Fault, shot time too short', class Mixing Head Warning, trigger "Mixinghead_MHControl3_DBW_6" bit 15
   15209: 'Mixinghead 03: Mixinghead collides when opening or closing', class Mixing Head Warning, trigger "Mixinghead_MHControl3_DBW_6" bit 0
   15210: 'Mixinghead 03: Runtime monitoring when locking mixing head', class Mixing Head Warning, trigger "Mixinghead_MHControl3_DBW_6" bit 1
   15211: 'Mixinghead 03: Runtime monitoring when unlocking mixing head', class Mixing Head Warning, trigger "Mixinghead_MHControl3_DBW_6" bit 2
   15212: 'Mixinghead 03:', class Mixing Head Warning, trigger "Mixinghead_MHControl3_DBW_6" bit 3
   15213: 'Mixinghead 03:', class Mixing Head Warning, trigger "Mixinghead_MHControl3_DBW_6" bit 4
   15214: 'Mixinghead 03:', class Mixing Head Warning, trigger "Mixinghead_MHControl3_DBW_6" bit 5
   15215: 'Mixinghead 03:', class Mixing Head Warning, trigger "Mixinghead_MHControl3_DBW_6" bit 6
   15216: 'Mixinghead 03: Component required in entry is not enabled at this mixing head', class Mixing Head Errors, trigger "Mixinghead_MHControl3_DBW_6" bit 7
   15217: 'Mixinghead 03: Cleaning piston: Moving out too slow', class Mixing Head Errors, trigger "Mixinghead_Cpiston3_DBW_38" bit 8
   15218: 'Mixinghead 03: Cleaning piston: Moving in too slow', class Mixing Head Errors, trigger "Mixinghead_Cpiston3_DBW_38" bit 9
   15219: 'Mixinghead 03: Cleaning piston: Proximity switch defect', class Mixing Head Errors, trigger "Mixinghead_Cpiston3_DBW_38" bit 10
   15220: 'Mixinghead 03: Cleaning piston: Leaves its home position in entry', class Mixing Head Errors, trigger "Mixinghead_Cpiston3_DBW_38" bit 11
   15221: 'Mixinghead 03: Cleaning piston: Not defined', class Mixing Head Warning, trigger "Mixinghead_Cpiston3_DBW_38" bit 12
   15222: 'Mixinghead 03: Cleaning piston:', class Mixing Head Warning, trigger "Mixinghead_Cpiston3_DBW_38" bit 13
   15223: 'Mixinghead 03: Cleaning piston:', class Mixing Head Warning, trigger "Mixinghead_Cpiston3_DBW_38" bit 14
   15224: 'Mixinghead 03: Cleaning piston:', class Mixing Head Warning, trigger "Mixinghead_Cpiston3_DBW_38" bit 15
   15225: 'Mixinghead 03: Cleaning piston: Controller at upper limit', class Mixing Head Warning, trigger "Mixinghead_Cpiston3_DBW_38" bit 0
   15226: 'Mixinghead 03: Cleaning piston: Controller at lower limit', class Mixing Head Warning, trigger "Mixinghead_Cpiston3_DBW_38" bit 1
   15227: 'Mixinghead 03: Cleaning piston:', class Mixing Head Warning, trigger "Mixinghead_Cpiston3_DBW_38" bit 2
   15228: 'Mixinghead 03: Cleaning piston: Front position not reached', class Mixing Head Warning, trigger "Mixinghead_Cpiston3_DBW_38" bit 3
   15229: 'Mixinghead 03: Cleaning piston: Rear position not reached', class Mixing Head Warning, trigger "Mixinghead_Cpiston3_DBW_38" bit 4
   15230: 'Mixinghead 03: Cleaning piston: Home position not reached', class Mixing Head Warning, trigger "Mixinghead_Cpiston3_DBW_38" bit 5
   15231: 'Mixinghead 03: Cleaning piston:', class Mixing Head Warning, trigger "Mixinghead_Cpiston3_DBW_38" bit 6
   15232: 'Mixinghead 03: Cleaning piston:', class Mixing Head Warning, trigger "Mixinghead_Cpiston3_DBW_38" bit 7
   15240: 'Mixinghead 03: Connection 01: Temperature recording: Measuring value outside measuring range', class Mixing Head Warning, trigger "Mixinghead_Temperature_MH3_Con1_DBW74" bit 8
   15241: 'Mixinghead 03: Connection 01: Temperature recording: Warning, value exceeded', class Mixing Head Warning, trigger "Mixinghead_Temperature_MH3_Con1_DBW74" bit 9
   15242: 'Mixinghead 03: Connection 01: Temperature recording: Warning, value undershot', class Mixing Head Warning, trigger "Mixinghead_Temperature_MH3_Con1_DBW74" bit 10
   15243: 'Mixinghead 03: Connection 01: Temperature recording: Fault, value exceeded', class Mixing Head Errors, trigger "Mixinghead_Temperature_MH3_Con1_DBW74" bit 11
   15244: 'Mixinghead 03: Connection 01: Temperature recording: Fault, value undershot', class Mixing Head Errors, trigger "Mixinghead_Temperature_MH3_Con1_DBW74" bit 12
   15245: 'Mixinghead 03: Connection 02: Temperature recording: Measuring value outside measuring range', class Mixing Head Warning, trigger "Mixinghead_Temperature_MH3_Con2_DBW108" bit 8
   15246: 'Mixinghead 03: Connection 02: Temperature recording: Warning, value exceeded', class Mixing Head Warning, trigger "Mixinghead_Temperature_MH3_Con2_DBW108" bit 9
   15247: 'Mixinghead 03: Connection 02: Temperature recording: Warning, value undershot', class Mixing Head Warning, trigger "Mixinghead_Temperature_MH3_Con2_DBW108" bit 10
   15248: 'Mixinghead 03: Connection 02: Temperature recording: Fault, value exceeded', class Mixing Head Errors, trigger "Mixinghead_Temperature_MH3_Con2_DBW108" bit 11
   15249: 'Mixinghead 03: Connection 02: Temperature recording: Fault, value undershot', class Mixing Head Errors, trigger "Mixinghead_Temperature_MH3_Con2_DBW108" bit 12
   15250: 'Mixinghead 03: Connection 03: Temperature recording: Measuring value outside measuring range', class Mixing Head Warning, trigger "Mixinghead_Temperature_MH3_Con3_DBW142" bit 8
   15251: 'Mixinghead 03: Connection 03: Temperature recording: Warning, value exceeded', class Mixing Head Warning, trigger "Mixinghead_Temperature_MH3_Con3_DBW142" bit 9
   15252: 'Mixinghead 03: Connection 03: Temperature recording: Warning, value undershot', class Mixing Head Warning, trigger "Mixinghead_Temperature_MH3_Con3_DBW142" bit 10
   15253: 'Mixinghead 03: Connection 03: Temperature recording: Fault, value exceeded', class Mixing Head Errors, trigger "Mixinghead_Temperature_MH3_Con3_DBW142" bit 11
   15254: 'Mixinghead 03: Connection 03: Temperature recording: Fault, value undershot', class Mixing Head Errors, trigger "Mixinghead_Temperature_MH3_Con3_DBW142" bit 12
   15255: 'Mixinghead 03: Connection 04: Temperature recording: Measuring value outside measuring range', class Mixing Head Warning, trigger "Mixinghead_Temperature_MH3_Con4_DBW176" bit 8
   15256: 'Mixinghead 03: Connection 04: Temperature recording: Warning, value exceeded', class Mixing Head Warning, trigger "Mixinghead_Temperature_MH3_Con4_DBW176" bit 9
   15257: 'Mixinghead 03: Connection 04: Temperature recording: Warning, value undershot', class Mixing Head Warning, trigger "Mixinghead_Temperature_MH3_Con4_DBW176" bit 10
   15258: 'Mixinghead 03: Connection 04: Temperature recording: Fault, value exceeded', class Mixing Head Errors, trigger "Mixinghead_Temperature_MH3_Con4_DBW176" bit 11
   15259: 'Mixinghead 03: Connection 04: Temperature recording: Fault, value undershot', class Mixing Head Errors, trigger "Mixinghead_Temperature_MH3_Con4_DBW176" bit 12
   15260: 'Mixinghead 03: Connection 05: Temperature recording: Measuring value outside measuring range', class Mixing Head Warning, trigger "Mixinghead_Temperature_MH3_Con5_DBW210" bit 8
   15261: 'Mixinghead 03: Connection 05: Temperature recording: Warning, value exceeded', class Mixing Head Warning, trigger "Mixinghead_Temperature_MH3_Con5_DBW210" bit 9
   15262: 'Mixinghead 03: Connection 05: Temperature recording: Warning, value undershot', class Mixing Head Warning, trigger "Mixinghead_Temperature_MH3_Con5_DBW210" bit 10
   15263: 'Mixinghead 03: Connection 05: Temperature recording: Fault, value exceeded', class Mixing Head Errors, trigger "Mixinghead_Temperature_MH3_Con5_DBW210" bit 11
   15264: 'Mixinghead 03: Connection 05: Temperature recording: Fault, value undershot', class Mixing Head Errors, trigger "Mixinghead_Temperature_MH3_Con5_DBW210" bit 12
   15265: 'Mixinghead 03: Connection 06: Temperature recording: Measuring value outside measuring range', class Mixing Head Warning, trigger "Mixinghead_Temperature_MH3_Con6_DBW244" bit 8
   15266: 'Mixinghead 03: Connection 06: Temperature recording: Warning, value exceeded', class Mixing Head Warning, trigger "Mixinghead_Temperature_MH3_Con6_DBW244" bit 9
   15267: 'Mixinghead 03: Connection 06: Temperature recording: Warning, value undershot', class Mixing Head Warning, trigger "Mixinghead_Temperature_MH3_Con6_DBW244" bit 10
   15268: 'Mixinghead 03: Connection 06: Temperature recording: Fault, value exceeded', class Mixing Head Errors, trigger "Mixinghead_Temperature_MH3_Con6_DBW244" bit 11
   15269: 'Mixinghead 03: Connection 06: Temperature recording: Fault, value undershot', class Mixing Head Errors, trigger "Mixinghead_Temperature_MH3_Con6_DBW244" bit 12
   15270: 'Mixinghead 03: Connection 01: Pressure recording: Measuring value outside measuring range', class Mixing Head Warning, trigger "Mixinghead_Pressure_MH3_Con1_DBW278" bit 8
   15271: 'Mixinghead 03: Connection 01: Pressure recording: Warning, value exceeded', class Mixing Head Warning, trigger "Mixinghead_Pressure_MH3_Con1_DBW278" bit 9
   15272: 'Mixinghead 03: Connection 01: Pressure recording: Warning, value undershot', class Mixing Head Warning, trigger "Mixinghead_Pressure_MH3_Con1_DBW278" bit 10
   15273: 'Mixinghead 03: Connection 01: Pressure recording: Fault, value exceeded', class Mixing Head Errors, trigger "Mixinghead_Pressure_MH3_Con1_DBW278" bit 11
   15274: 'Mixinghead 03: Connection 01: Pressure recording: Fault, value undershot', class Mixing Head Errors, trigger "Mixinghead_Pressure_MH3_Con1_DBW278" bit 12
   15275: 'Mixinghead 03: Connection 02: Pressure recording: Measuring value outside measuring range', class Mixing Head Warning, trigger "Mixinghead_Pressure_MH3_Con2_DBW312" bit 8
   15276: 'Mixinghead 03: Connection 02: Pressure recording: Warning, value exceeded', class Mixing Head Warning, trigger "Mixinghead_Pressure_MH3_Con2_DBW312" bit 9
   15277: 'Mixinghead 03: Connection 02: Pressure recording: Warning, value undershot', class Mixing Head Warning, trigger "Mixinghead_Pressure_MH3_Con2_DBW312" bit 10
   15278: 'Mixinghead 03: Connection 02: Pressure recording: Fault, value exceeded', class Mixing Head Errors, trigger "Mixinghead_Pressure_MH3_Con2_DBW312" bit 11
   15279: 'Mixinghead 03: Connection 02: Pressure recording: Fault, value undershot', class Mixing Head Errors, trigger "Mixinghead_Pressure_MH3_Con2_DBW312" bit 12
   15280: 'Mixinghead 03: Connection 03: Pressure recording: Measuring value outside measuring range', class Mixing Head Warning, trigger "Mixinghead_Pressure_MH3_Con3_DBW346" bit 8
   15281: 'Mixinghead 03: Connection 03: Pressure recording: Warning, value exceeded', class Mixing Head Warning, trigger "Mixinghead_Pressure_MH3_Con3_DBW346" bit 9
   15282: 'Mixinghead 03: Connection 03: Pressure recording: Warning, value undershot', class Mixing Head Warning, trigger "Mixinghead_Pressure_MH3_Con3_DBW346" bit 10
   15283: 'Mixinghead 03: Connection 03: Pressure recording: Fault, value exceeded', class Mixing Head Errors, trigger "Mixinghead_Pressure_MH3_Con3_DBW346" bit 11
   15284: 'Mixinghead 03: Connection 03: Pressure recording: Fault, value undershot', class Mixing Head Errors, trigger "Mixinghead_Pressure_MH3_Con3_DBW346" bit 12
   15285: 'Mixinghead 03: Connection 04: Pressure recording: Measuring value outside measuring range', class Mixing Head Warning, trigger "Mixinghead_Pressure_MH3_Con4_DBW380" bit 8
   15286: 'Mixinghead 03: Connection 04: Pressure recording: Warning, value exceeded', class Mixing Head Warning, trigger "Mixinghead_Pressure_MH3_Con4_DBW380" bit 9
   15287: 'Mixinghead 03: Connection 04: Pressure recording: Warning, value undershot', class Mixing Head Warning, trigger "Mixinghead_Pressure_MH3_Con4_DBW380" bit 10
   15288: 'Mixinghead 03: Connection 04: Pressure recording: Fault, value exceeded', class Mixing Head Errors, trigger "Mixinghead_Pressure_MH3_Con4_DBW380" bit 11
   15289: 'Mixinghead 03: Connection 04: Pressure recording: Fault, value undershot', class Mixing Head Errors, trigger "Mixinghead_Pressure_MH3_Con4_DBW380" bit 12
   15290: 'Mixinghead 03: Connection 05: Pressure recording: Measuring value outside measuring range', class Mixing Head Warning, trigger "Mixinghead_Pressure_MH3_Con5_DBW414" bit 8
   15291: 'Mixinghead 03: Connection 05: Pressure recording: Warning, value exceeded', class Mixing Head Warning, trigger "Mixinghead_Pressure_MH3_Con5_DBW414" bit 9
   15292: 'Mixinghead 03: Connection 05: Pressure recording: Warning, value undershot', class Mixing Head Warning, trigger "Mixinghead_Pressure_MH3_Con5_DBW414" bit 10
   15293: 'Mixinghead 03: Connection 05: Pressure recording: Fault, value exceeded', class Mixing Head Errors, trigger "Mixinghead_Pressure_MH3_Con5_DBW414" bit 11
   15294: 'Mixinghead 03: Connection 05: Pressure recording: Fault, value undershot', class Mixing Head Errors, trigger "Mixinghead_Pressure_MH3_Con5_DBW414" bit 12
   15295: 'Mixinghead 03: Connection 06: Pressure recording: Measuring value outside measuring range', class Mixing Head Warning, trigger "Mixinghead_Pressure_MH3_Con6_DBW448" bit 8
   15296: 'Mixinghead 03: Connection 06: Pressure recording: Warning, value exceeded', class Mixing Head Warning, trigger "Mixinghead_Pressure_MH3_Con6_DBW448" bit 1
   15297: 'Mixinghead 03: Connection 06: Pressure recording: Warning, value undershot', class Mixing Head Warning, trigger "Mixinghead_Pressure_MH3_Con6_DBW448" bit 2
   15298: 'Mixinghead 03: Connection 06: Pressure recording: Fault, value exceeded', class Mixing Head Errors, trigger "Mixinghead_Pressure_MH3_Con6_DBW448" bit 3
   15299: 'Mixinghead 03: Connection 06: Pressure recording: Fault, value undershot', class Mixing Head Errors, trigger "Mixinghead_Pressure_MH3_Con6_DBW448" bit 4
   15301: 'Mixinghead 04: Mixinghead does not open', class Mixing Head Errors, trigger "Mixinghead_MHControl4_DBW_8" bit 8
   15302: 'Mixinghead 04: Mixinghead does not close', class Mixing Head Errors, trigger "Mixinghead_MHControl4_DBW_8" bit 9
   15303: 'Mixinghead 04: Entry cancelled', class Mixing Head Warning, trigger "Mixinghead_MHControl4_DBW_8" bit 10
   15304: 'Mixinghead 04: Mixinghead open without activation', class Mixing Head Errors, trigger "Mixinghead_MHControl4_DBW_8" bit 11
   15305: 'Mixinghead 04: Mixinghead close during entry', class Mixing Head Warning, trigger "Mixinghead_MHControl4_DBW_8" bit 12
   15306: 'Mixinghead 04: Warning, shot time too short', class Mixing Head Warning, trigger "Mixinghead_MHControl4_DBW_8" bit 13
   15307: 'Mixinghead 04: Warning , shot time too long', class Mixing Head Warning, trigger "Mixinghead_MHControl4_DBW_8" bit 14
   15308: 'Mixinghead 04: Fault, shot time too short', class Mixing Head Warning, trigger "Mixinghead_MHControl4_DBW_8" bit 15
   15309: 'Mixinghead 04: Mixinghead collides when opening or closing', class Mixing Head Warning, trigger "Mixinghead_MHControl4_DBW_8" bit 0
   15310: 'Mixinghead 04: Runtime monitoring when locking mixing head', class Mixing Head Warning, trigger "Mixinghead_MHControl4_DBW_8" bit 1
   15311: 'Mixinghead 04: Runtime monitoring when unlocking mixing head', class Mixing Head Warning, trigger "Mixinghead_MHControl4_DBW_8" bit 2
   15312: 'Mixinghead 04:', class Mixing Head Warning, trigger "Mixinghead_MHControl4_DBW_8" bit 3
   15313: 'Mixinghead 04:', class Mixing Head Warning, trigger "Mixinghead_MHControl4_DBW_8" bit 4
   15314: 'Mixinghead 04:', class Mixing Head Warning, trigger "Mixinghead_MHControl4_DBW_8" bit 5
   15315: 'Mixinghead 04:', class Mixing Head Warning, trigger "Mixinghead_MHControl4_DBW_8" bit 6
   15316: 'Mixinghead 04: Component required in entry is not enabled at this mixing head', class Mixing Head Errors, trigger "Mixinghead_MHControl4_DBW_8" bit 7
   15317: 'Mixinghead 04: Cleaning piston: Moving out too slow', class Mixing Head Errors, trigger "Mixinghead_Cpiston4_DBW_40" bit 8
   15318: 'Mixinghead 04: Cleaning piston: Moving in too slow', class Mixing Head Errors, trigger "Mixinghead_Cpiston4_DBW_40" bit 9
   15319: 'Mixinghead 04: Cleaning piston: Proximity switch defect', class Mixing Head Errors, trigger "Mixinghead_Cpiston4_DBW_40" bit 10
   15320: 'Mixinghead 04: Cleaning piston: Leaves its home position in entry', class Mixing Head Errors, trigger "Mixinghead_Cpiston4_DBW_40" bit 11
   15321: 'Mixinghead 04: Cleaning piston: Not defined', class Mixing Head Warning, trigger "Mixinghead_Cpiston4_DBW_40" bit 12
   15322: 'Mixinghead 04: Cleaning piston:', class Mixing Head Warning, trigger "Mixinghead_Cpiston4_DBW_40" bit 13
   15323: 'Mixinghead 04: Cleaning piston:', class Mixing Head Warning, trigger "Mixinghead_Cpiston4_DBW_40" bit 14
   15324: 'Mixinghead 04: Cleaning piston:', class Mixing Head Warning, trigger "Mixinghead_Cpiston4_DBW_40" bit 15
   15325: 'Mixinghead 04: Cleaning piston: Controller at upper limit', class Mixing Head Warning, trigger "Mixinghead_Cpiston4_DBW_40" bit 0
   15326: 'Mixinghead 04: Cleaning piston: Controller at lower limit', class Mixing Head Warning, trigger "Mixinghead_Cpiston4_DBW_40" bit 1
   15327: 'Mixinghead 04: Cleaning piston:', class Mixing Head Warning, trigger "Mixinghead_Cpiston4_DBW_40" bit 2